(* Logix 5000 project; controller TemplateV1R0 vendor 1 type 14 code 222 rev 33.11; software revision 33.00; part 3 of 5 *)
(* tags used below, declared in another part *)
   Sts_Show_HMIControls : BOOL;   // 0 = dont show 1 = Show controls
   T_Switch_Time : TIMER[2];   // timer for valve to move from open to close or the otherway around
   ons_reset : BOOL;   // prevent continious reset
   T_Mem_Valve : TIMER[2];
(* Valve_V2, continued *)

ROUTINE Prescan   (* structured text *)
   ////////////////////////////////////////////////////////////
   //   Copyright (c)
   //------------------------------------------------------------
   //   Routine: Prescan
   //   Author: WPI\tom.reit
   //   Created: 28-11-2022
   //------------------------------------------------------------
   //   Description:
   //
   //
   //   History:
   //
   ////////////////////////////////////////////////////////////
   if T_Switch_Time[0].PRE = 0 then T_Switch_Time[0].PRE:=500; end_if;
   if T_Switch_Time[1].PRE = 0 then T_Switch_Time[1].PRE:=500; end_if;
   T_Mem_Valve[0].PRE:=50;
   T_Mem_Valve[1].PRE:=50;
   
   Sts_Show_HMIControls :=0;
   
END_ROUTINE
END_ADD_ON_INSTRUCTION

ADD_ON_INSTRUCTION WaterCircuit   (* revision 1.1, vendor WPI, ExecutePrescan *)
// Closed water circuit based on Micro820
VAR_INPUT
   Reset : BOOL; {required}   // Reset WTU C1&C2 on falling edge of reset signal
   Select_Mode : BOOL; {visible}   // 1 = Automatic 0 = Manual
   Start : BOOL; {visible}   // 0 = OFF 1 = ON
END_VAR
VAR_OUTPUT
   Temperature : REAL; {access Read Only, visible}   // Actual Temperature (c)
END_VAR
VAR_INPUT
   PID_CycleTime : DINT; {required}   // Cycle time for SSR
   PID_Kc : LREAL; {required}   // Proportional and Integral are dependent on this gain. (>= 0.0001). Increasing Kc improves response time but also increases overshoot and oscillation of the PID.
   PID_Ti : LREAL; {required}   // Time integral constant in seconds (>= 0.0001). Increasing Ti decreases the overshoot and oscillation of the PID.
   PID_Td : LREAL; {required}   // Time derivative constant in seconds (>= 0.0). When Td equals 0, there is no derivative action and PID becomes a PI controller. Increasing Td reduces the overshot and removes the oscillation of the PID controller.
   PID_FC : LREAL; {required}   // Filter constant (>= 0.0). Recommended range for FC is 0 to 20. Increasing FC smooths the response of the PID controller.
   PID_Setpoint : LREAL; {visible}   // Setpoint temperature (c)
END_VAR
VAR_OUTPUT
   PID_OUTPUT : REAL; {access Read Only, visible}   // Output PID controller (%)
END_VAR
VAR_INPUT
   PID_HandValue : LREAL; {visible}   // handvalue in % of time
   ManualStart_CP : BOOL; {visible}   // 0 = OFF 1 = ON
   ManualStart_HE : BOOL; {visible}   // 0 = OFF 1 = ON
   ManualStart_V1 : BOOL; {visible}   // 0 = OFF 1 = ON
   ManualStart_V2 : BOOL; {visible}   // 0 = OFF 1 = ON
END_VAR
VAR_OUTPUT
   ALARM_CommunicationFaulted : BOOL; {access Read Only, visible}   // Communication faulted, check IP address in MSG instruction
   ALARM_Active : BOOL; {access Read Only, visible}   // Alarm is active, outputs will NOT be activated on WTU
   ALARM_PressureFaulted : BOOL; {access Read Only, visible}   // Filling faulted
   ALARM_Overload_CirculationPump : BOOL; {access Read Only, visible}   // Overload_CirculationPump
   ALARM_Overload_Heatingelement : BOOL; {access Read Only, visible}   // Overload_Heatingelment
   ALARM_Max_TemperatureSwitch : BOOL; {access Read Only, visible}   // Max TemperatureSwitch
   ALARM_TemperatureSensorLost : BOOL; {access Read Only, visible}   // cable disconnected temperature sensor
   Sts_Communication_OK : BOOL; {access Read Only, visible}   // Communication is OK to micro820
   Sts_CirculationPump : BOOL; {access Read Only, visible}   // Status Circulationpump output
   Sts_HeatingElement : BOOL; {access Read Only, visible}   // Status Heating element output
   Sts_SolidstateRelais : BOOL; {access Read Only, visible}   // Status SSR output
   Sts_CoolingValve : BOOL; {access Read Only, visible}   // Status Cooling Valve output
   Sts_FillingValve : BOOL; {access Read Only, visible}   // Status Filling Valve output
END_VAR
VAR_IN_OUT
   Read_Element : LREAL[40]; {required}   // Dataholder
   Msg_Read : MESSAGE; {required}   // Message to read object
   Write_Element : LREAL[40]; {required}   // Dataholder
   Msg_Write : MESSAGE; {required}   // Message to read object
END_VAR
VAR_INPUT
   Enable_Communication : BOOL; {visible}   // set to true if messages can be send to micro820
   cnf_Select_Circuit : USINT;   // assign AOI to watercircuit based on: 1 = C1 2 = C2
END_VAR
VAR_OUTPUT
   HMI_Color : DINT; {access Read Only}   // 0 = off 1 = auto turned on 2 = manual control 3= no communication
END_VAR
VAR
   RefreshRate : FBD_TIMER; {access None}   // refreshrate timer
   wrk_conversion : DINT[20]; {access None}   // conversion tag to go from LREAL to DINT
   i : SINT; {access None}   // local index num
   InputStatus : DINT; {access None}   // InputStatus from Micro820
        .12   // spare
        .0   // _IO_EM_DI_00
        .1   // _IO_EM_DI_01
        .10   // _IO_EM_DI_10
        .11   // _IO_EM_DI_11
        .13   // spare
        .14   // spare
        .15   // spare
        .16   // spare
        .17   // spare
        .18   // spare
        .19   // spare
        .2   // _IO_EM_DI_02
        .20   // spare
        .21   // spare
        .22   // spare
        .23   // spare
        .24   // spare
        .25   // spare
        .26   // spare
        .27   // spare
        .28   // spare
        .29   // spare
        .3   // _IO_EM_DI_03
        .30   // spare
        .31   // spare
        .4   // _IO_EM_DI_04
        .5   // _IO_EM_DI_05
        .6   // _IO_EM_DI_06
        .7   // _IO_EM_DI_07
        .8   // _IO_EM_DI_08
        .9   // _IO_EM_DI_09
   TagName : STRING; {access Read Only}   // Contains tag name based on addon name
   HMI_Trend_MaxValue : DINT; {access Read Only}   // Trend for HMI
   HMI_Trend_MinValue : DINT; {access Read Only}   // HMI_Trend_MinValue
END_VAR

ROUTINE Logic   (* structured text *)
// Closed water circuit based on Micro820
   ////////////////////////////////////////////////////////////
   //   Copyright (c)
   //------------------------------------------------------------
   //   Routine: WaterCircuit - Logic
   //   Author: WPI\tom.reit
   //   Created: 13-3-2023
   //------------------------------------------------------------
   //   Description:
   //           Closed water circuit based on Micro820
   //
   //
   //   History:
   //
   ////////////////////////////////////////////////////////////
   RefreshRate.EN:=1;
   RefreshRate.PRE:=50;
   RefreshRate.TimerEnable:=1;
   RefreshRate.Reset:=RefreshRate.DN;
   TONR(RefreshRate);
   if RefreshRate.DN then
   	MSG(Msg_Read);																	// Message to read object. CIP datatable read.
   	MSG(Msg_Write);																	// Message to Write object. CIP datatable write.
   end_if;
   #region Message OK
   	if Msg_Read.DN AND Msg_Write.DN then
   		Sts_Communication_OK:=1;
   	end_if;
   	if NOT Enable_Communication then
   		Sts_Communication_OK:=0;
   	end_if;
   #endregion
   #region Message timeout/faulted
   	if Msg_Read.ER OR Msg_Write.ER then
   		ALARM_CommunicationFaulted:=1;
   		Sts_Communication_OK:=0;
   	else
   		ALARM_CommunicationFaulted:=0;
   	end_if;
   	if Reset AND (Msg_Read.ER OR Msg_Write.ER)  then
   		Msg_Read.Flags			:=0;	// reset Message instruction
   		Msg_Write.Flags			:=0;	// reset Message instruction
   	end_if;
   #endregion
   for i := 0 to 19 do
   	wrk_conversion[i]:=0;// clear old data
   end_for;
   wrk_conversion[0].0			:=		Reset;						// Micro820 tag: HMI_I_Reset
   
   /* Prevent wrong user input */
   if cnf_Select_Circuit > 2 then cnf_Select_Circuit:=2; end_if;
   if cnf_Select_Circuit < 1 then cnf_Select_Circuit:=1; end_if;
   
   #region Convert IO from Micro820 to local
   	wrk_conversion[18]				:=		Read_Element[18];	// InputStatus
   	InputStatus						:= 		wrk_conversion[18];
   	wrk_conversion[19]				:=		Read_Element[19];	// OutputStatus
   #endregion
   if Enable_Communication then
   	#region data
   		#region Convert InputData to LREAL
   			wrk_conversion[1].0			:=		Select_Mode;				// Micro820 tag: HMI_I_C1_Select_Mode
   			wrk_conversion[2].0			:=		Start;					// Micro820 tag: HMI_I_StartC1
   			wrk_conversion[3].0			:=		ManualStart_CP;			// Micro820 tag: HMI_I_C1_ManualStart_CP
   			wrk_conversion[4].0			:=		ManualStart_HE;			// Micro820 tag: HMI_I_C1_ManualStart_HE
   			wrk_conversion[5].0			:=		ManualStart_V1;			// Micro820 tag: HMI_I_C1_ManualStart_V1
   			wrk_conversion[6].0			:=		ManualStart_V2;			// Micro820 tag: HMI_I_C1_ManualStart_V2
   			// IS ALLREADY A REAL, DOESNT NEED CONVERSION! 					// Micro820 tag: HMI_I_C1_Kc
   			// IS ALLREADY A REAL, DOESNT NEED CONVERSION! 					// Micro820 tag: HMI_I_C1_Ti
   			// IS ALLREADY A REAL, DOESNT NEED CONVERSION! 					// Micro820 tag: HMI_I_C1_Td
   			// IS ALLREADY A REAL, DOESNT NEED CONVERSION! 					// Micro820 tag: HMI_I_C1_FC
   			// IS ALLREADY A REAL, DOESNT NEED CONVERSION! 					// Micro820 tag: HMI_I_C1_PID_Setpoint
   			// IS ALLREADY A REAL, DOESNT NEED CONVERSION!					// Micro820 tag: HMI_I_C1_PID_HandValue
   			wrk_conversion[13]			:=		PID_CycleTime;			// Micro820 tag: HMI_I_C1_PID_CycleTime
   		/* set data for micro820 tag */
   		Write_Element[00]:=wrk_conversion[00];
   		Write_Element[01]:=wrk_conversion[01];
   		Write_Element[02]:=wrk_conversion[02];
   		Write_Element[03]:=wrk_conversion[03];
   		Write_Element[04]:=wrk_conversion[04];
   		Write_Element[05]:=wrk_conversion[05];
   		Write_Element[06]:=wrk_conversion[06];
   		Write_Element[07]:=PID_Kc;
   		Write_Element[08]:=PID_Ti;
   		Write_Element[09]:=PID_Td;
   		Write_Element[10]:=PID_FC;
   		Write_Element[11]:=PID_Setpoint;
   		Write_Element[12]:=PID_HandValue;
   		Write_Element[13]:=wrk_conversion[13];
   		#endregion
   		#region OutputData
   			Temperature						:=		Read_Element[0];
   			PID_OUTPUT						:=		Read_Element[1];
   
   			wrk_conversion[2]				:=		Read_Element[2];
   			ALARM_PressureFaulted			:=		wrk_conversion[2].0;
   
   			wrk_conversion[3]				:=		Read_Element[3];
   			ALARM_Overload_CirculationPump	:=		wrk_conversion[3].0;
   
   			wrk_conversion[4]				:=		Read_Element[4];
   			ALARM_Overload_Heatingelement	:=		wrk_conversion[4].0;
   
   			wrk_conversion[5]				:=		Read_Element[5];
   			ALARM_Max_TemperatureSwitch		:=		wrk_conversion[5].0;
   
   			wrk_conversion[6]				:=		Read_Element[6];
   			ALARM_TemperatureSensorLost		:=		wrk_conversion[6].0;
   
   			wrk_conversion[7]				:=		Read_Element[7];
   			ALARM_Active					:=		wrk_conversion[7].0;
   
   			if cnf_Select_Circuit = 1 then
   				Sts_CirculationPump				:=		wrk_conversion[19].0;
   				Sts_HeatingElement				:=		wrk_conversion[19].1;
   				Sts_SolidstateRelais			:=		wrk_conversion[19].2;
   				Sts_CoolingValve				:=		wrk_conversion[19].3;
   				Sts_FillingValve				:=		wrk_conversion[19].4;
   			elsif cnf_Select_Circuit = 2 then
   				Sts_CirculationPump				:=		wrk_conversion[19].5;
   				Sts_HeatingElement				:=		wrk_conversion[19].6;
   				Sts_SolidstateRelais			:=		wrk_conversion[19].7;
   				Sts_CoolingValve				:=		wrk_conversion[19].8;
   				Sts_FillingValve				:=		wrk_conversion[19].9;
   			end_if;
   		#endregion
   	#endregion
   end_if;
   #region HMI data visuals
   	if 	(Enable_Communication AND Sts_Communication_OK )  AND Select_Mode AND NOT Start then			// Auto - Turned off
   		HMI_Color:=0;
   	elsif (Enable_Communication AND Sts_Communication_OK )  AND Select_Mode AND Start then				// Auto - Turned on
   		HMI_Color:=1;
   	elsif (Enable_Communication AND Sts_Communication_OK )  AND NOT Select_Mode  then					// Manual - controlled manually
   		HMI_Color:=2;
   	elsif (Enable_Communication AND NOT Sts_Communication_OK ) then										// No connection
   		HMI_Color:=0;
   	elsif NOT Enable_Communication then																	// No connection
   		HMI_Color:=3;
   	end_if;
   	gsv(AddOnInstructionDefinition,THIS,Name,TagName);
   	if HMI_Trend_MaxValue=0 AND HMI_Trend_MinValue=0 then HMI_Trend_MaxValue:=100;HMI_Trend_MinValue:=0; end_if;
   #endregion
END_ROUTINE

ROUTINE Prescan   (* structured text *)
   ////////////////////////////////////////////////////////////
   //   Copyright (c)
   //------------------------------------------------------------
   //   Routine: Prescan
   //   Author: WPI\tom.reit
   //   Created: 15-3-2023
   //------------------------------------------------------------
   //   Description:
   //
   //
   //   History:
   //
   ////////////////////////////////////////////////////////////
   Enable_Communication:=1;
END_ROUTINE
END_ADD_ON_INSTRUCTION

VAR_GLOBAL   (* controller tags *)
   SafetyZone1_Unit1_Reset : BOOL;
END_VAR

PROGRAM MainProgram   (* main routine MainRoutine *)

ROUTINE MainRoutine   (* ladder *)
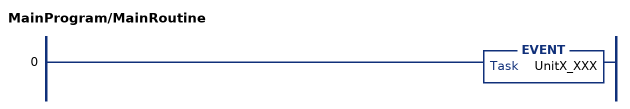
   0: EVENT(UnitX_XXX);
END_ROUTINE
END_PROGRAM

PROGRAM SafetyProgram   (* main routine MainRoutine, safety *)

ROUTINE MainRoutine   (* ladder *)
END_ROUTINE
END_PROGRAM

PROGRAM UnitX_EMXXX   (* main routine Main *)
VAR
   Alarm : AlarmGenerator[10] := ([1].Alarm_ID := 1, [2].Alarm_ID := 2, [3].Alarm_ID := 3, [4].Alarm_ID := 4, [5].Alarm_ID := 5, [6].Alarm_ID := 6, [7].Alarm_ID := 7, [8].Alarm_ID := 8, [9].Alarm_ID := 9);
   AlarmText : STRING[10] := ([1] := '| Unit4_Batter_EM01_Depositor | X-axis faulted | ', [2] := '| Unit4_Batter_EM01_Depositor | Y-axis faulted |', [3] := '| Unit4_Batter_EM01_Depositor | Z-axis faulted |', [4] := '| Unit4_Batter_EM01_Depositor | Manifold ColorInjected-axis faulted |', [5] := '| Unit4_Batter_EM01_Depositor | No Color Manifold-axis faulted |', [6] := '| Unit4_Batter_EM01_Depositor | Overload servo drives |', [7] := '| Unit4_Batter_EM01_Depositor | X,Y,Z Motion faulted |', [8] := '| Unit4_Batter_EM01_Depositor | Manifold Motion faulted |', [9] := '| Unit1_Sander_EM01_Elende |');
   wrk_mode_Select : DINT := 1;   // mode select for case
   wrk_StartNum : DINT := 100;   // StartStateModelNum
   wrk_state_Select : DINT := 9;   // select correct prog
END_VAR

ROUTINE _EP_00_Selector   (* structured text *)
   ////////////////////////////////////////////////////////////
   //   Copyright (c)
   //------------------------------------------------------------
   //   Routine: _EP_00_Selector
   //   Author: WPI\tom.reit
   //   Created: 11-11-2022
   //------------------------------------------------------------
   //   Description:
   //
   //
   //   History:
   //
   ////////////////////////////////////////////////////////////
   if 		Unit.Sts_Production 	then	wrk_mode_Select:=1;
   elsif 	Unit.Sts_Maintenance 	then	wrk_mode_Select:=2;
   elsif 	Unit.Sts_Manual 		then	wrk_mode_Select:=3;
   elsif 	Unit.Sts_Cleaning 		then	wrk_mode_Select:=4;
   elsif 	Unit.Sts_MES 			then	wrk_mode_Select:=5;
   elsif 	Unit.Sts_SemiAutomatic 	then	wrk_mode_Select:=6;
   end_if;
   #region Set case state non active states
   	if 		Unit.Sts_Aborted 		then	wrk_state_Select:=9;
   	elsif 	Unit.Sts_Stopped		then	wrk_state_Select:=2;
   	elsif   Unit.Sts_Idle			then	wrk_state_Select:=4;
   	elsif 	Unit.Sts_Execute		then	wrk_state_Select:=6;
   	elsif 	Unit.Sts_Held			then	wrk_state_Select:=11;
   	elsif 	Unit.Sts_Suspended		then	wrk_state_Select:=5;
   	elsif   Unit.Sts_Complete		then	wrk_state_Select:=17;
   	end_if;
   #endregion
   #region Set case state
   	if 		Unit.Sts_Production AND Unit.Sts_Aborting 		then	wrk_state_Select:=8;
   	elsif 	Unit.Sts_Production AND Unit.Sts_Clearing		then	wrk_state_Select:=1;
   	elsif 	Unit.Sts_Production AND Unit.Sts_Stopping		then	wrk_state_Select:=7;
   	elsif 	Unit.Sts_Production	AND Unit.Sts_Resetting		then	wrk_state_Select:=15;
   	elsif 	Unit.Sts_Production AND Unit.Sts_Starting		then	wrk_state_Select:=3;
   	elsif 	Unit.Sts_Production AND Unit.Sts_Holding		then	wrk_state_Select:=10;
   	elsif 	Unit.Sts_Production AND Unit.Sts_Unholding		then	wrk_state_Select:=12;
   	elsif 	Unit.Sts_Production AND Unit.Sts_Suspending		then	wrk_state_Select:=13;
   	elsif 	Unit.Sts_Production AND Unit.Sts_Unsuspending	then	wrk_state_Select:=14;
   	elsif 	Unit.Sts_Production AND Unit.Sts_Completing		then	wrk_state_Select:=16;
   	end_if;
   #endregion
   #region Set case state
   	if 		Unit.Sts_Maintenance AND Unit.Sts_Aborting 		then	wrk_state_Select:=8;
   	elsif 	Unit.Sts_Maintenance AND Unit.Sts_Clearing		then	wrk_state_Select:=1;
   	elsif 	Unit.Sts_Maintenance AND Unit.Sts_Stopping		then	wrk_state_Select:=7;
   	elsif 	Unit.Sts_Maintenance AND Unit.Sts_Resetting		then	wrk_state_Select:=15;
   	elsif 	Unit.Sts_Maintenance AND Unit.Sts_Starting		then	wrk_state_Select:=3;
   	elsif 	Unit.Sts_Maintenance AND Unit.Sts_Holding		then	wrk_state_Select:=10;
   	elsif 	Unit.Sts_Maintenance AND Unit.Sts_Unholding		then	wrk_state_Select:=12;
   	elsif 	Unit.Sts_Maintenance AND Unit.Sts_Suspending	then	wrk_state_Select:=13;
   	elsif 	Unit.Sts_Maintenance AND Unit.Sts_Unsuspending	then	wrk_state_Select:=14;
   	elsif 	Unit.Sts_Maintenance AND Unit.Sts_Completing	then	wrk_state_Select:=16;
   	end_if;
   #endregion
   #region Set case state
   	if 		Unit.Sts_Manual AND Unit.Sts_Aborting 		then	wrk_state_Select:=8;
   	elsif 	Unit.Sts_Manual AND Unit.Sts_Clearing		then	wrk_state_Select:=1;
   	elsif 	Unit.Sts_Manual AND Unit.Sts_Stopping		then	wrk_state_Select:=7;
   	elsif 	Unit.Sts_Manual	AND Unit.Sts_Resetting		then	wrk_state_Select:=15;
   	elsif 	Unit.Sts_Manual AND Unit.Sts_Starting		then	wrk_state_Select:=3;
   	elsif 	Unit.Sts_Manual AND Unit.Sts_Holding		then	wrk_state_Select:=10;
   	elsif 	Unit.Sts_Manual AND Unit.Sts_Unholding		then	wrk_state_Select:=12;
   	elsif 	Unit.Sts_Manual AND Unit.Sts_Suspending		then	wrk_state_Select:=13;
   	elsif 	Unit.Sts_Manual AND Unit.Sts_Unsuspending	then	wrk_state_Select:=14;
   	elsif 	Unit.Sts_Manual AND Unit.Sts_Completing		then	wrk_state_Select:=16;
   	end_if;
   #endregion
   #region Set case state
   	if 		Unit.Sts_Cleaning AND Unit.Sts_Aborting 	then	wrk_state_Select:=8;
   	elsif 	Unit.Sts_Cleaning AND Unit.Sts_Clearing		then	wrk_state_Select:=1;
   	elsif 	Unit.Sts_Cleaning AND Unit.Sts_Stopping		then	wrk_state_Select:=7;
   	elsif 	Unit.Sts_Cleaning AND Unit.Sts_Resetting	then	wrk_state_Select:=15;
   	elsif 	Unit.Sts_Cleaning AND Unit.Sts_Starting		then	wrk_state_Select:=3;
   	elsif 	Unit.Sts_Cleaning AND Unit.Sts_Holding		then	wrk_state_Select:=10;
   	elsif 	Unit.Sts_Cleaning AND Unit.Sts_Unholding	then	wrk_state_Select:=12;
   	elsif 	Unit.Sts_Cleaning AND Unit.Sts_Suspending	then	wrk_state_Select:=13;
   	elsif 	Unit.Sts_Cleaning AND Unit.Sts_Unsuspending	then	wrk_state_Select:=14;
   	elsif 	Unit.Sts_Cleaning AND Unit.Sts_Completing	then	wrk_state_Select:=16;
   	end_if;
   #endregion
   #region Set case state
   	if 		Unit.Sts_MES AND Unit.Sts_Aborting 		then	wrk_state_Select:=8;
   	elsif 	Unit.Sts_MES AND Unit.Sts_Clearing		then	wrk_state_Select:=1;
   	elsif 	Unit.Sts_MES AND Unit.Sts_Stopping		then	wrk_state_Select:=7;
   	elsif 	Unit.Sts_MES AND Unit.Sts_Resetting		then	wrk_state_Select:=15;
   	elsif 	Unit.Sts_MES AND Unit.Sts_Starting		then	wrk_state_Select:=3;
   	elsif 	Unit.Sts_MES AND Unit.Sts_Holding		then	wrk_state_Select:=10;
   	elsif 	Unit.Sts_MES AND Unit.Sts_Unholding		then	wrk_state_Select:=12;
   	elsif 	Unit.Sts_MES AND Unit.Sts_Suspending	then	wrk_state_Select:=13;
   	elsif 	Unit.Sts_MES AND Unit.Sts_Unsuspending	then	wrk_state_Select:=14;
   	elsif 	Unit.Sts_MES AND Unit.Sts_Completing	then	wrk_state_Select:=16;
   	end_if;
   #endregion
   #region Set case state
   	if 		Unit.Sts_SemiAutomatic AND Unit.Sts_Aborting 		then	wrk_state_Select:=8;
   	elsif 	Unit.Sts_SemiAutomatic AND Unit.Sts_Clearing		then	wrk_state_Select:=1;
   	elsif 	Unit.Sts_SemiAutomatic AND Unit.Sts_Stopping		then	wrk_state_Select:=7;
   	elsif 	Unit.Sts_SemiAutomatic	AND Unit.Sts_Resetting		then	wrk_state_Select:=15;
   	elsif 	Unit.Sts_SemiAutomatic AND Unit.Sts_Starting		then	wrk_state_Select:=3;
   	elsif 	Unit.Sts_SemiAutomatic AND Unit.Sts_Holding			then	wrk_state_Select:=10;
   	elsif 	Unit.Sts_SemiAutomatic AND Unit.Sts_Unholding		then	wrk_state_Select:=12;
   	elsif 	Unit.Sts_SemiAutomatic AND Unit.Sts_Suspending		then	wrk_state_Select:=13;
   	elsif 	Unit.Sts_SemiAutomatic AND Unit.Sts_Unsuspending	then	wrk_state_Select:=14;
   	elsif 	Unit.Sts_SemiAutomatic AND Unit.Sts_Completing		then	wrk_state_Select:=16;
   	end_if;
   #endregion
   
   
   EquipmentModule.Request_SC.ons_Reset.InputBit:=Unit.Sts_MachineFaulted OR EquipmentModule.Reset_Signal;
   OSRI(EquipmentModule.Request_SC.ons_Reset);
   if EquipmentModule.Request_SC.ons_Reset.OutputBit then
   	EquipmentModule.EP_SEQ.Holding		:=0;
   	EquipmentModule.EP_SEQ.Starting		:=0;
   	EquipmentModule.EP_SEQ.Suspending	:=0;
   	EquipmentModule.EP_SEQ.Unholding	:=0;
   	EquipmentModule.EP_SEQ.Unsuspending	:=0;
   end_if;
   
   if EquipmentModule.Force_Stop OR EquipmentModule.Force_Abort then EquipmentModule.Faulted:=1; else EquipmentModule.Faulted:=0; end_if;
   case wrk_mode_Select of
   	1:																	/* Production(automatic) */
   		wrk_StartNum:=100;
   		case wrk_state_Select of
   			1: 	JSR(_EP_01_Clearing); 		if EquipmentModule.EP_SEQ.Clearing		=0 then EquipmentModule.EP_SEQ.Clearing		:=wrk_StartNum; 	end_if;
   			3: 	JSR(_EP_03_Starting);		if EquipmentModule.EP_SEQ.Starting		=0 then EquipmentModule.EP_SEQ.Starting		:=wrk_StartNum; 	end_if;
   			6: 	JSR(_EP_06_Execute);
   			7: 	JSR(_EP_07_Stopping);		if EquipmentModule.EP_SEQ.Stopping		=0 then EquipmentModule.EP_SEQ.Stopping		:=wrk_StartNum; 	end_if;
   			8: 	JSR(_EP_08_Aborting); 		if EquipmentModule.EP_SEQ.Aborting		=0 then EquipmentModule.EP_SEQ.Aborting		:=wrk_StartNum; 	end_if;
   			10: JSR(_EP_10_Holding);		if EquipmentModule.EP_SEQ.Holding		=0 then EquipmentModule.EP_SEQ.Holding		:=wrk_StartNum; 	end_if;
   			12:	JSR(_EP_12_Unholding);		if EquipmentModule.EP_SEQ.Unholding		=0 then EquipmentModule.EP_SEQ.Unholding	:=wrk_StartNum; 	end_if;
   			13:	JSR(_EP_13_Suspending);		if EquipmentModule.EP_SEQ.Suspending	=0 then EquipmentModule.EP_SEQ.Suspending	:=wrk_StartNum; 	end_if;
   			14:	JSR(_EP_14_Unsuspending);	if EquipmentModule.EP_SEQ.Unsuspending	=0 then EquipmentModule.EP_SEQ.Unsuspending	:=wrk_StartNum; 	end_if;
   			15:	JSR(_EP_15_Resetting);		if EquipmentModule.EP_SEQ.Resetting		=0 then EquipmentModule.EP_SEQ.Resetting	:=wrk_StartNum; 	end_if;
   			16:	JSR(_EP_16_Completing);		if EquipmentModule.EP_SEQ.Completing	=0 then EquipmentModule.EP_SEQ.Completing	:=wrk_StartNum; 	end_if;
   			else
   		end_case;
   	2:																	/* Maintenance */
   		wrk_StartNum:=200;
   		case wrk_state_Select of
   			1: 	JSR(_EP_01_Clearing); 		if EquipmentModule.EP_SEQ.Clearing		=0 then EquipmentModule.EP_SEQ.Clearing		:=wrk_StartNum; 	end_if;
   			3: 	JSR(_EP_03_Starting);		if EquipmentModule.EP_SEQ.Starting		=0 then EquipmentModule.EP_SEQ.Starting		:=wrk_StartNum; 	end_if;
   			6: 	JSR(_EP_06_Execute);
   			7: 	JSR(_EP_07_Stopping);		if EquipmentModule.EP_SEQ.Stopping		=0 then EquipmentModule.EP_SEQ.Stopping		:=wrk_StartNum; 	end_if;
   			8: 	JSR(_EP_08_Aborting); 		if EquipmentModule.EP_SEQ.Aborting		=0 then EquipmentModule.EP_SEQ.Aborting		:=wrk_StartNum; 	end_if;
   			10: JSR(_EP_10_Holding);		if EquipmentModule.EP_SEQ.Holding		=0 then EquipmentModule.EP_SEQ.Holding		:=wrk_StartNum; 	end_if;
   			12:	JSR(_EP_12_Unholding);		if EquipmentModule.EP_SEQ.Unholding		=0 then EquipmentModule.EP_SEQ.Unholding	:=wrk_StartNum; 	end_if;
   			13:	JSR(_EP_13_Suspending);		if EquipmentModule.EP_SEQ.Suspending	=0 then EquipmentModule.EP_SEQ.Suspending	:=wrk_StartNum; 	end_if;
   			14:	JSR(_EP_14_Unsuspending);	if EquipmentModule.EP_SEQ.Unsuspending	=0 then EquipmentModule.EP_SEQ.Unsuspending	:=wrk_StartNum; 	end_if;
   			15:	JSR(_EP_15_Resetting);		if EquipmentModule.EP_SEQ.Resetting		=0 then EquipmentModule.EP_SEQ.Resetting	:=wrk_StartNum; 	end_if;
   			16:	JSR(_EP_16_Completing);		if EquipmentModule.EP_SEQ.Completing	=0 then EquipmentModule.EP_SEQ.Completing	:=wrk_StartNum; 	end_if;
   			else
   		end_case;
   	3:																	/* Manual */
   		wrk_StartNum:=300;
   		case wrk_state_Select of
   			1: 	JSR(_EP_01_Clearing); 		if EquipmentModule.EP_SEQ.Clearing		=0 then EquipmentModule.EP_SEQ.Clearing		:=wrk_StartNum; 	end_if;
   			3: 	JSR(_EP_03_Starting);		if EquipmentModule.EP_SEQ.Starting		=0 then EquipmentModule.EP_SEQ.Starting		:=wrk_StartNum; 	end_if;
   			6: 	JSR(_EP_06_Execute);
   			7: 	JSR(_EP_07_Stopping);		if EquipmentModule.EP_SEQ.Stopping		=0 then EquipmentModule.EP_SEQ.Stopping		:=wrk_StartNum; 	end_if;
   			8: 	JSR(_EP_08_Aborting); 		if EquipmentModule.EP_SEQ.Aborting		=0 then EquipmentModule.EP_SEQ.Aborting		:=wrk_StartNum; 	end_if;
   			10: JSR(_EP_10_Holding);		if EquipmentModule.EP_SEQ.Holding		=0 then EquipmentModule.EP_SEQ.Holding		:=wrk_StartNum; 	end_if;
   			12:	JSR(_EP_12_Unholding);		if EquipmentModule.EP_SEQ.Unholding		=0 then EquipmentModule.EP_SEQ.Unholding	:=wrk_StartNum; 	end_if;
   			13:	JSR(_EP_13_Suspending);		if EquipmentModule.EP_SEQ.Suspending	=0 then EquipmentModule.EP_SEQ.Suspending	:=wrk_StartNum; 	end_if;
   			14:	JSR(_EP_14_Unsuspending);	if EquipmentModule.EP_SEQ.Unsuspending	=0 then EquipmentModule.EP_SEQ.Unsuspending	:=wrk_StartNum; 	end_if;
   			15:	JSR(_EP_15_Resetting);		if EquipmentModule.EP_SEQ.Resetting		=0 then EquipmentModule.EP_SEQ.Resetting	:=wrk_StartNum; 	end_if;
   			16:	JSR(_EP_16_Completing);		if EquipmentModule.EP_SEQ.Completing	=0 then EquipmentModule.EP_SEQ.Completing	:=wrk_StartNum; 	end_if;
   			else
   		end_case;
   	4:																	/* Cleaning */
   		wrk_StartNum:=400;
   		case wrk_state_Select of
   			1: 	JSR(_EP_01_Clearing); 		if EquipmentModule.EP_SEQ.Clearing		=0 then EquipmentModule.EP_SEQ.Clearing		:=wrk_StartNum; 	end_if;
   			3: 	JSR(_EP_03_Starting);		if EquipmentModule.EP_SEQ.Starting		=0 then EquipmentModule.EP_SEQ.Starting		:=wrk_StartNum; 	end_if;
   			6: 	JSR(_EP_06_Execute);
   			7: 	JSR(_EP_07_Stopping);		if EquipmentModule.EP_SEQ.Stopping		=0 then EquipmentModule.EP_SEQ.Stopping		:=wrk_StartNum; 	end_if;
   			8: 	JSR(_EP_08_Aborting); 		if EquipmentModule.EP_SEQ.Aborting		=0 then EquipmentModule.EP_SEQ.Aborting		:=wrk_StartNum; 	end_if;
   			10: JSR(_EP_10_Holding);		if EquipmentModule.EP_SEQ.Holding		=0 then EquipmentModule.EP_SEQ.Holding		:=wrk_StartNum; 	end_if;
   			12:	JSR(_EP_12_Unholding);		if EquipmentModule.EP_SEQ.Unholding		=0 then EquipmentModule.EP_SEQ.Unholding	:=wrk_StartNum; 	end_if;
   			13:	JSR(_EP_13_Suspending);		if EquipmentModule.EP_SEQ.Suspending	=0 then EquipmentModule.EP_SEQ.Suspending	:=wrk_StartNum; 	end_if;
   			14:	JSR(_EP_14_Unsuspending);	if EquipmentModule.EP_SEQ.Unsuspending	=0 then EquipmentModule.EP_SEQ.Unsuspending	:=wrk_StartNum; 	end_if;
   			15:	JSR(_EP_15_Resetting);		if EquipmentModule.EP_SEQ.Resetting		=0 then EquipmentModule.EP_SEQ.Resetting	:=wrk_StartNum; 	end_if;
   			16:	JSR(_EP_16_Completing);		if EquipmentModule.EP_SEQ.Completing	=0 then EquipmentModule.EP_SEQ.Completing	:=wrk_StartNum; 	end_if;
   			else
   		end_case;
   	5:																	/* MES */
   		wrk_StartNum:=500;
   		case wrk_state_Select of
   			1: 	JSR(_EP_01_Clearing); 		if EquipmentModule.EP_SEQ.Clearing		=0 then EquipmentModule.EP_SEQ.Clearing		:=wrk_StartNum; 	end_if;
   			3: 	JSR(_EP_03_Starting);		if EquipmentModule.EP_SEQ.Starting		=0 then EquipmentModule.EP_SEQ.Starting		:=wrk_StartNum; 	end_if;
   			6: 	JSR(_EP_06_Execute);
   			7: 	JSR(_EP_07_Stopping);		if EquipmentModule.EP_SEQ.Stopping		=0 then EquipmentModule.EP_SEQ.Stopping		:=wrk_StartNum; 	end_if;
   			8: 	JSR(_EP_08_Aborting); 		if EquipmentModule.EP_SEQ.Aborting		=0 then EquipmentModule.EP_SEQ.Aborting		:=wrk_StartNum; 	end_if;
   			10: JSR(_EP_10_Holding);		if EquipmentModule.EP_SEQ.Holding		=0 then EquipmentModule.EP_SEQ.Holding		:=wrk_StartNum; 	end_if;
   			12:	JSR(_EP_12_Unholding);		if EquipmentModule.EP_SEQ.Unholding		=0 then EquipmentModule.EP_SEQ.Unholding	:=wrk_StartNum; 	end_if;
   			13:	JSR(_EP_13_Suspending);		if EquipmentModule.EP_SEQ.Suspending	=0 then EquipmentModule.EP_SEQ.Suspending	:=wrk_StartNum; 	end_if;
   			14:	JSR(_EP_14_Unsuspending);	if EquipmentModule.EP_SEQ.Unsuspending	=0 then EquipmentModule.EP_SEQ.Unsuspending	:=wrk_StartNum; 	end_if;
   			15:	JSR(_EP_15_Resetting);		if EquipmentModule.EP_SEQ.Resetting		=0 then EquipmentModule.EP_SEQ.Resetting	:=wrk_StartNum; 	end_if;
   			16:	JSR(_EP_16_Completing);		if EquipmentModule.EP_SEQ.Completing	=0 then EquipmentModule.EP_SEQ.Completing	:=wrk_StartNum; 	end_if;
   			else
   		end_case;
   	6:																	/* semiautomatic */
   		wrk_StartNum:=600;
   		case wrk_state_Select of
   			1: 	JSR(_EP_01_Clearing); 		if EquipmentModule.EP_SEQ.Clearing		=0 then EquipmentModule.EP_SEQ.Clearing		:=wrk_StartNum; 	end_if;
   			3: 	JSR(_EP_03_Starting);		if EquipmentModule.EP_SEQ.Starting		=0 then EquipmentModule.EP_SEQ.Starting		:=wrk_StartNum; 	end_if;
   			6: 	JSR(_EP_06_Execute);
   			7: 	JSR(_EP_07_Stopping);		if EquipmentModule.EP_SEQ.Stopping		=0 then EquipmentModule.EP_SEQ.Stopping		:=wrk_StartNum; 	end_if;
   			8: 	JSR(_EP_08_Aborting); 		if EquipmentModule.EP_SEQ.Aborting		=0 then EquipmentModule.EP_SEQ.Aborting		:=wrk_StartNum; 	end_if;
   			10: JSR(_EP_10_Holding);		if EquipmentModule.EP_SEQ.Holding		=0 then EquipmentModule.EP_SEQ.Holding		:=wrk_StartNum; 	end_if;
   			12:	JSR(_EP_12_Unholding);		if EquipmentModule.EP_SEQ.Unholding		=0 then EquipmentModule.EP_SEQ.Unholding	:=wrk_StartNum; 	end_if;
   			13:	JSR(_EP_13_Suspending);		if EquipmentModule.EP_SEQ.Suspending	=0 then EquipmentModule.EP_SEQ.Suspending	:=wrk_StartNum; 	end_if;
   			14:	JSR(_EP_14_Unsuspending);	if EquipmentModule.EP_SEQ.Unsuspending	=0 then EquipmentModule.EP_SEQ.Unsuspending	:=wrk_StartNum; 	end_if;
   			15:	JSR(_EP_15_Resetting);		if EquipmentModule.EP_SEQ.Resetting		=0 then EquipmentModule.EP_SEQ.Resetting	:=wrk_StartNum; 	end_if;
   			16:	JSR(_EP_16_Completing);		if EquipmentModule.EP_SEQ.Completing	=0 then EquipmentModule.EP_SEQ.Completing	:=wrk_StartNum; 	end_if;
   			else
   		end_case;
   	else
   		wrk_mode_Select:=1;
   end_case;
   
   													/* Reset SC signals once machine is next state */
   if Unit.Sts_Aborted 	AND EquipmentModule.Request_SC.Aborting_to_Aborted 		then EquipmentModule.Request_SC.Aborting_to_Aborted			:=0; 	end_if;
   if Unit.Sts_Complete 	AND EquipmentModule.Request_SC.Completing_to_Completed 	then EquipmentModule.Request_SC.Completing_to_Completed		:=0; 	end_if;
   if Unit.Sts_Execute 	AND EquipmentModule.Request_SC.Starting_to_Execute 		then EquipmentModule.Request_SC.Starting_to_Execute			:=0; 	end_if;
   if Unit.Sts_Complete 	AND EquipmentModule.Request_SC.Execute_to_Completing 	then EquipmentModule.Request_SC.Execute_to_Completing		:=0; 	end_if;
   if Unit.Sts_Execute 	AND EquipmentModule.Request_SC.Unholding_to_Execute 	then EquipmentModule.Request_SC.Unholding_to_Execute		:=0; 	end_if;
   if Unit.Sts_Execute 	AND EquipmentModule.Request_SC.Unsuspending_to_Execute 	then EquipmentModule.Request_SC.Unsuspending_to_Execute		:=0; 	end_if;
   if Unit.Sts_Held 		AND EquipmentModule.Request_SC.Holding_to_Held 			then EquipmentModule.Request_SC.Holding_to_Held				:=0; 	end_if;
   if Unit.Sts_Idle 		AND EquipmentModule.Request_SC.Resetting_to_Idle 		then EquipmentModule.Request_SC.Resetting_to_Idle			:=0; 	end_if;
   if Unit.Sts_Stopped 	AND EquipmentModule.Request_SC.Clearing_to_Stopped 		then EquipmentModule.Request_SC.Clearing_to_Stopped 		:=0; 	end_if;
   if Unit.Sts_Stopped 	AND EquipmentModule.Request_SC.Stopping_to_Stopped 		then EquipmentModule.Request_SC.Stopping_to_Stopped			:=0; 	end_if;
   if Unit.Sts_Suspended 	AND EquipmentModule.Request_SC.Suspending_to_Suspended 	then EquipmentModule.Request_SC.Suspending_to_Suspended		:=0; 	end_if;
   
   													/* Reset SEQ once machine is next state */
   if Unit.Sts_Aborted 	AND		EquipmentModule.EP_SEQ.Aborting<>0		then EquipmentModule.EP_SEQ.Aborting	:=0; end_if;
   if Unit.Sts_Stopped 	AND		EquipmentModule.EP_SEQ.Clearing<>0		then EquipmentModule.EP_SEQ.Clearing	:=0; end_if;
   if Unit.Sts_Stopped 	AND		EquipmentModule.EP_SEQ.Stopping<>0		then EquipmentModule.EP_SEQ.Stopping	:=0; end_if;
   if Unit.Sts_Idle 		AND		EquipmentModule.EP_SEQ.Resetting<>0		then EquipmentModule.EP_SEQ.Resetting	:=0; end_if;
   if Unit.Sts_Execute 	AND		EquipmentModule.EP_SEQ.Starting<>0		then EquipmentModule.EP_SEQ.Starting	:=0; end_if;
   if Unit.Sts_Execute 	AND		EquipmentModule.EP_SEQ.Unholding<>0		then EquipmentModule.EP_SEQ.Unholding	:=0; end_if;
   if Unit.Sts_Execute 	AND		EquipmentModule.EP_SEQ.Unsuspending<>0	then EquipmentModule.EP_SEQ.Unsuspending:=0; end_if;
   if Unit.Sts_Complete 	AND		EquipmentModule.EP_SEQ.Completing<>0	then EquipmentModule.EP_SEQ.Completing	:=0; end_if;
   if Unit.Sts_Held 		AND		EquipmentModule.EP_SEQ.Holding<>0		then EquipmentModule.EP_SEQ.Holding		:=0; end_if;
   if Unit.Sts_Suspended	AND		EquipmentModule.EP_SEQ.Suspending<>0	then EquipmentModule.EP_SEQ.Suspending	:=0; end_if;
   
   
   
   
   
   #region AlarmFeedback to Unit
   	Alarm[1].Alarm_ID:=1;
   	Alarm[2].Alarm_ID:=2;
   	Alarm[3].Alarm_ID:=3;
   	Alarm[4].Alarm_ID:=4;
   	Alarm[5].Alarm_ID:=5;
   	Alarm[6].Alarm_ID:=6;
   	Alarm[7].Alarm_ID:=7;
   	Alarm[8].Alarm_ID:=8;
   	Alarm[9].Alarm_ID:=9;
   	AlarmGenerator(Alarm[1],EquipmentModule,AlarmText[1]);
   	AlarmGenerator(Alarm[2],EquipmentModule,AlarmText[2]);
   	AlarmGenerator(Alarm[3],EquipmentModule,AlarmText[3]);
   	AlarmGenerator(Alarm[4],EquipmentModule,AlarmText[4]);
   	AlarmGenerator(Alarm[5],EquipmentModule,AlarmText[5]);
   	AlarmGenerator(Alarm[6],EquipmentModule,AlarmText[6]);
   	AlarmGenerator(Alarm[7],EquipmentModule,AlarmText[7]);
   	AlarmGenerator(Alarm[8],EquipmentModule,AlarmText[8]);
   	AlarmGenerator(Alarm[9],EquipmentModule,AlarmText[9]);
   #endregion
END_ROUTINE

ROUTINE _EP_01_Clearing   (* ladder *)
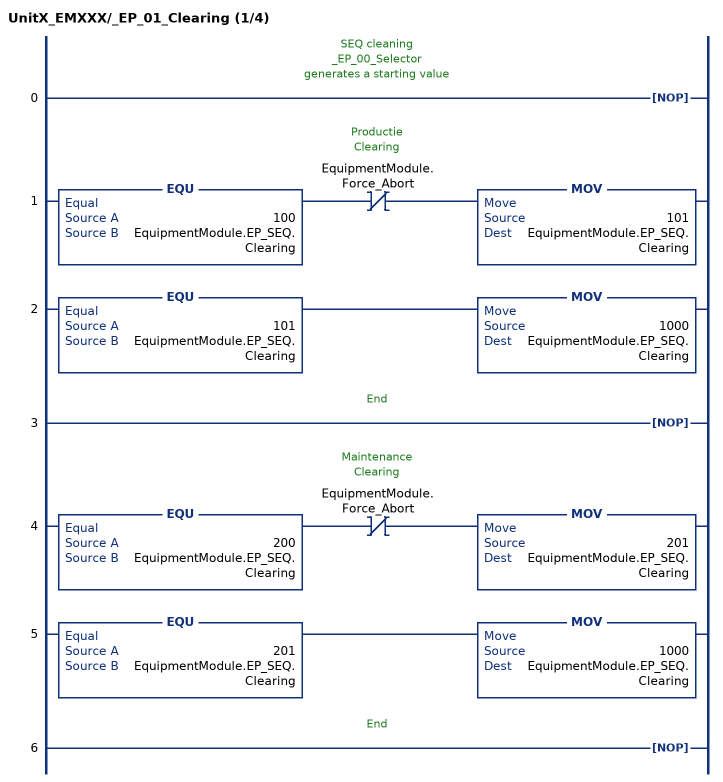
   // SEQ cleaning
   // _EP_00_Selector
   // generates a starting value
   0: NOP();
   // Productie
   // Clearing
   1: EQU(100,EquipmentModule.EP_SEQ.Clearing)XIO(EquipmentModule.Force_Abort)MOV(101,EquipmentModule.EP_SEQ.Clearing);
   2: EQU(101,EquipmentModule.EP_SEQ.Clearing)MOV(1000,EquipmentModule.EP_SEQ.Clearing);
   // End
   3: NOP();
   // Maintenance
   // Clearing
   4: EQU(200,EquipmentModule.EP_SEQ.Clearing)XIO(EquipmentModule.Force_Abort)MOV(201,EquipmentModule.EP_SEQ.Clearing);
   5: EQU(201,EquipmentModule.EP_SEQ.Clearing)MOV(1000,EquipmentModule.EP_SEQ.Clearing);
   // End
   6: NOP();
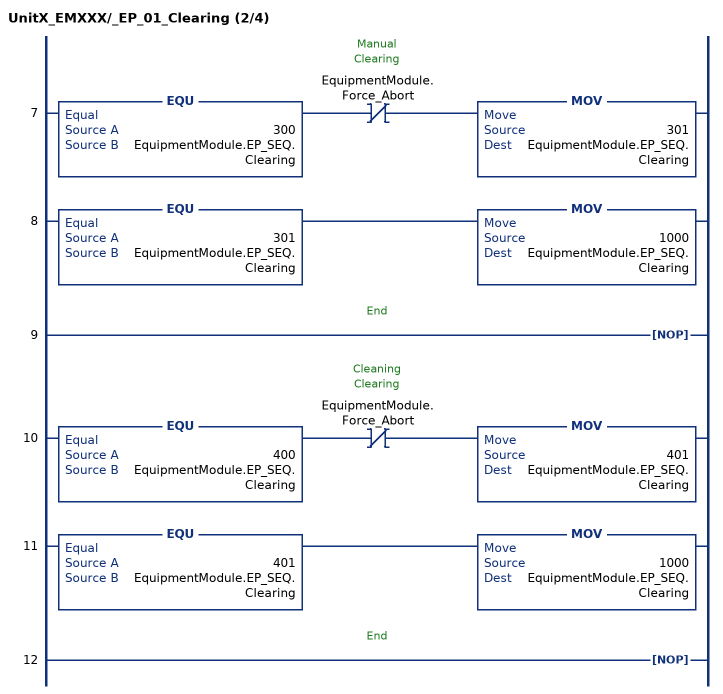
   // Manual
   // Clearing
   7: EQU(300,EquipmentModule.EP_SEQ.Clearing)XIO(EquipmentModule.Force_Abort)MOV(301,EquipmentModule.EP_SEQ.Clearing);
   8: EQU(301,EquipmentModule.EP_SEQ.Clearing)MOV(1000,EquipmentModule.EP_SEQ.Clearing);
   // End
   9: NOP();
   // Cleaning
   // Clearing
   10: EQU(400,EquipmentModule.EP_SEQ.Clearing)XIO(EquipmentModule.Force_Abort)MOV(401,EquipmentModule.EP_SEQ.Clearing);
   11: EQU(401,EquipmentModule.EP_SEQ.Clearing)MOV(1000,EquipmentModule.EP_SEQ.Clearing);
   // End
   12: NOP();
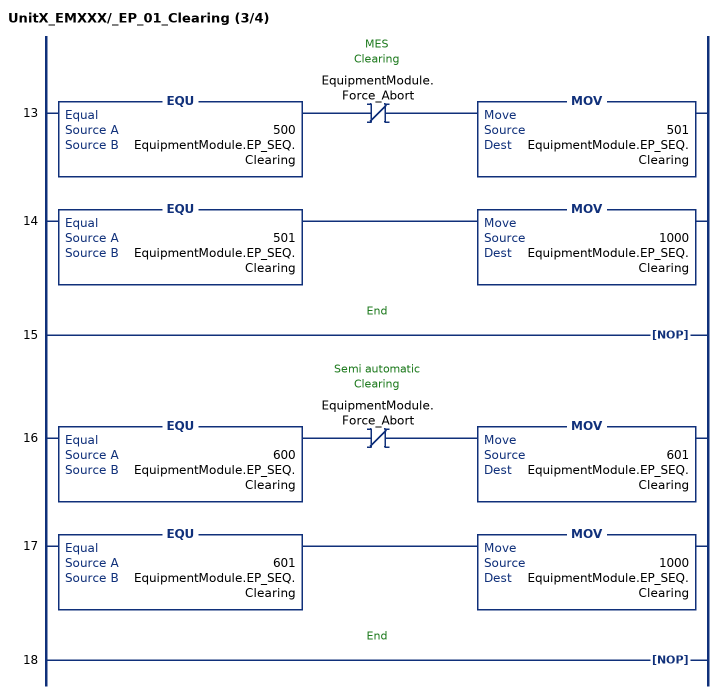
   // MES
   // Clearing
   13: EQU(500,EquipmentModule.EP_SEQ.Clearing)XIO(EquipmentModule.Force_Abort)MOV(501,EquipmentModule.EP_SEQ.Clearing);
   14: EQU(501,EquipmentModule.EP_SEQ.Clearing)MOV(1000,EquipmentModule.EP_SEQ.Clearing);
   // End
   15: NOP();
   // Semi automatic
   // Clearing
   16: EQU(600,EquipmentModule.EP_SEQ.Clearing)XIO(EquipmentModule.Force_Abort)MOV(601,EquipmentModule.EP_SEQ.Clearing);
   17: EQU(601,EquipmentModule.EP_SEQ.Clearing)MOV(1000,EquipmentModule.EP_SEQ.Clearing);
   // End
   18: NOP();
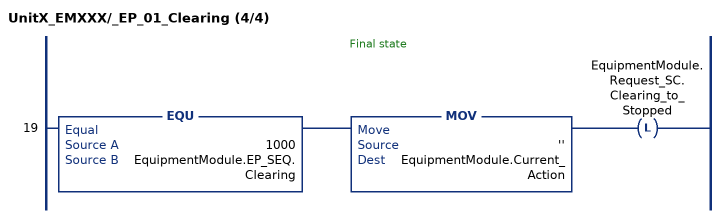
   // Final state
   19: EQU(1000,EquipmentModule.EP_SEQ.Clearing)MOV('',EquipmentModule.Current_Action)OTL(EquipmentModule.Request_SC.Clearing_to_Stopped);
END_ROUTINE

ROUTINE _EP_03_Starting   (* ladder *)
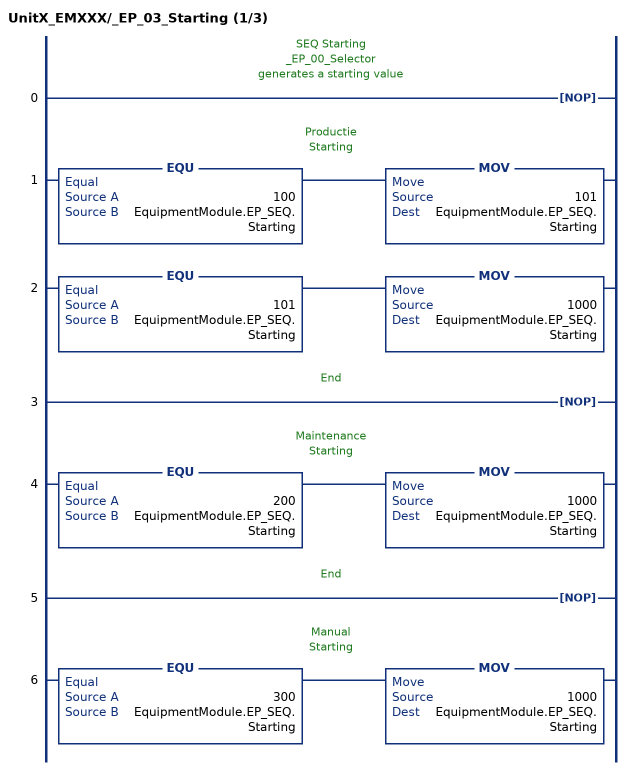
   // SEQ Starting
   // _EP_00_Selector
   // generates a starting value
   0: NOP();
   // Productie
   // Starting
   1: EQU(100,EquipmentModule.EP_SEQ.Starting)MOV(101,EquipmentModule.EP_SEQ.Starting);
   2: EQU(101,EquipmentModule.EP_SEQ.Starting)MOV(1000,EquipmentModule.EP_SEQ.Starting);
   // End
   3: NOP();
   // Maintenance
   // Starting
   4: EQU(200,EquipmentModule.EP_SEQ.Starting)MOV(1000,EquipmentModule.EP_SEQ.Starting);
   // End
   5: NOP();
   // Manual
   // Starting
   6: EQU(300,EquipmentModule.EP_SEQ.Starting)MOV(1000,EquipmentModule.EP_SEQ.Starting);
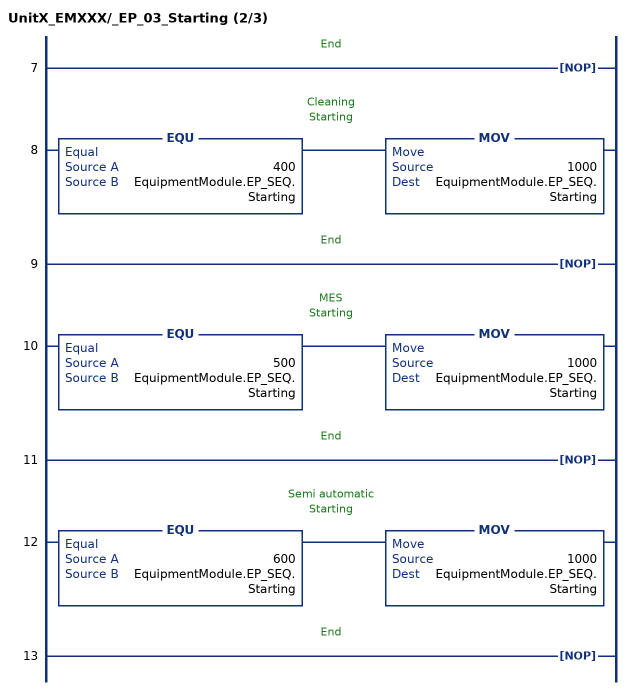
   // End
   7: NOP();
   // Cleaning
   // Starting
   8: EQU(400,EquipmentModule.EP_SEQ.Starting)MOV(1000,EquipmentModule.EP_SEQ.Starting);
   // End
   9: NOP();
   // MES
   // Starting
   10: EQU(500,EquipmentModule.EP_SEQ.Starting)MOV(1000,EquipmentModule.EP_SEQ.Starting);
   // End
   11: NOP();
   // Semi automatic
   // Starting
   12: EQU(600,EquipmentModule.EP_SEQ.Starting)MOV(1000,EquipmentModule.EP_SEQ.Starting);
   // End
   13: NOP();
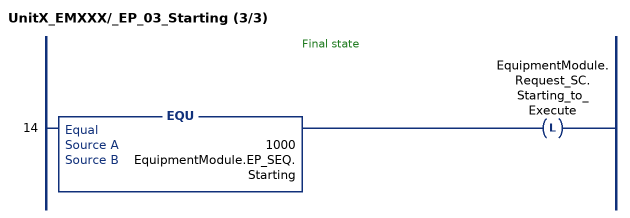
   // Final state
   14: EQU(1000,EquipmentModule.EP_SEQ.Starting)OTL(EquipmentModule.Request_SC.Starting_to_Execute);
END_ROUTINE

ROUTINE _EP_06_Execute   (* ladder *)
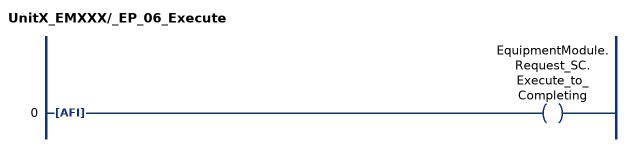
   0: AFI()OTE(EquipmentModule.Request_SC.Execute_to_Completing);
END_ROUTINE

ROUTINE _EP_07_Stopping   (* ladder *)
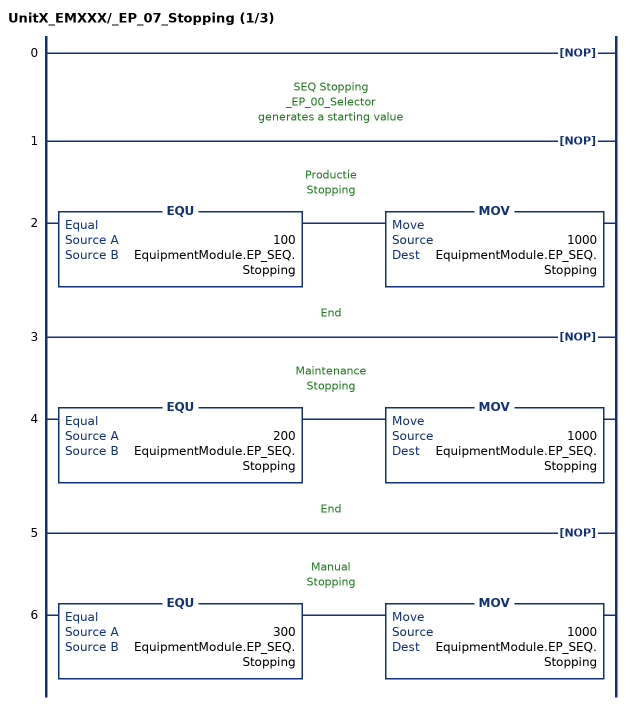
   0: NOP();
   // SEQ Stopping
   // _EP_00_Selector
   // generates a starting value
   1: NOP();
   // Productie
   // Stopping
   2: EQU(100,EquipmentModule.EP_SEQ.Stopping)MOV(1000,EquipmentModule.EP_SEQ.Stopping);
   // End
   3: NOP();
   // Maintenance
   // Stopping
   4: EQU(200,EquipmentModule.EP_SEQ.Stopping)MOV(1000,EquipmentModule.EP_SEQ.Stopping);
   // End
   5: NOP();
   // Manual
   // Stopping
   6: EQU(300,EquipmentModule.EP_SEQ.Stopping)MOV(1000,EquipmentModule.EP_SEQ.Stopping);
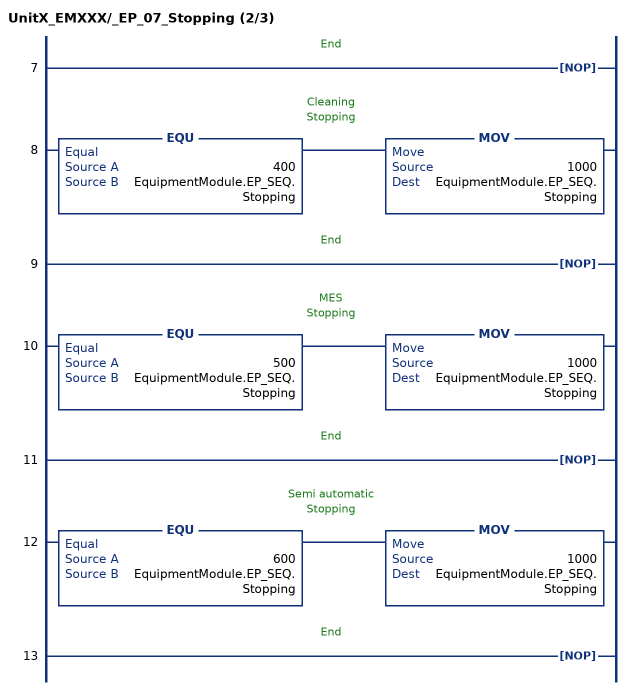
   // End
   7: NOP();
   // Cleaning
   // Stopping
   8: EQU(400,EquipmentModule.EP_SEQ.Stopping)MOV(1000,EquipmentModule.EP_SEQ.Stopping);
   // End
   9: NOP();
   // MES
   // Stopping
   10: EQU(500,EquipmentModule.EP_SEQ.Stopping)MOV(1000,EquipmentModule.EP_SEQ.Stopping);
   // End
   11: NOP();
   // Semi automatic
   // Stopping
   12: EQU(600,EquipmentModule.EP_SEQ.Stopping)MOV(1000,EquipmentModule.EP_SEQ.Stopping);
   // End
   13: NOP();
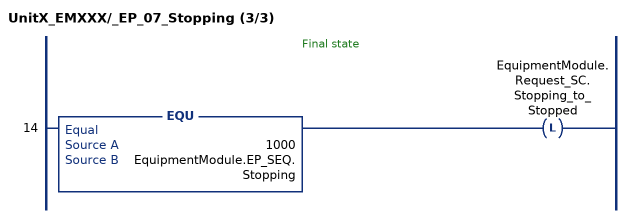
   // Final state
   14: EQU(1000,EquipmentModule.EP_SEQ.Stopping)OTL(EquipmentModule.Request_SC.Stopping_to_Stopped);
END_ROUTINE

ROUTINE _EP_08_Aborting   (* ladder *)
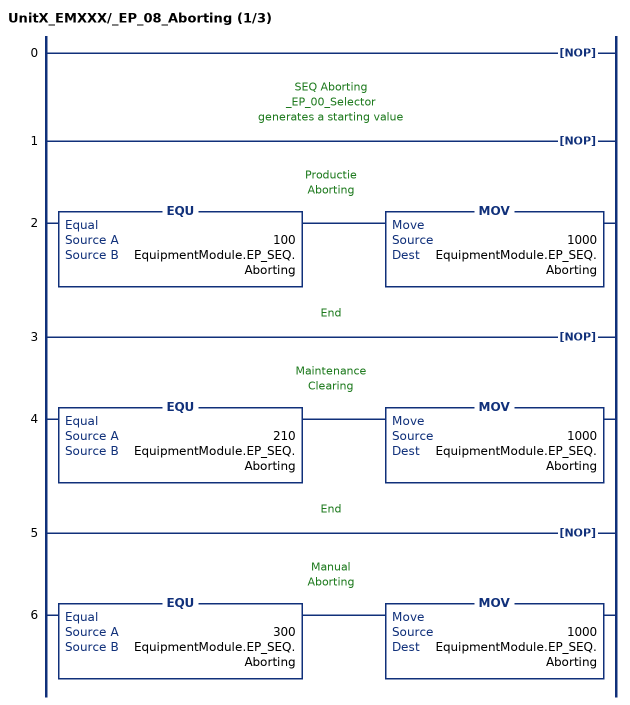
   0: NOP();
   // SEQ Aborting
   // _EP_00_Selector
   // generates a starting value
   1: NOP();
   // Productie
   // Aborting
   2: EQU(100,EquipmentModule.EP_SEQ.Aborting)MOV(1000,EquipmentModule.EP_SEQ.Aborting);
   // End
   3: NOP();
   // Maintenance
   // Clearing
   4: EQU(210,EquipmentModule.EP_SEQ.Aborting)MOV(1000,EquipmentModule.EP_SEQ.Aborting);
   // End
   5: NOP();
   // Manual
   // Aborting
   6: EQU(300,EquipmentModule.EP_SEQ.Aborting)MOV(1000,EquipmentModule.EP_SEQ.Aborting);
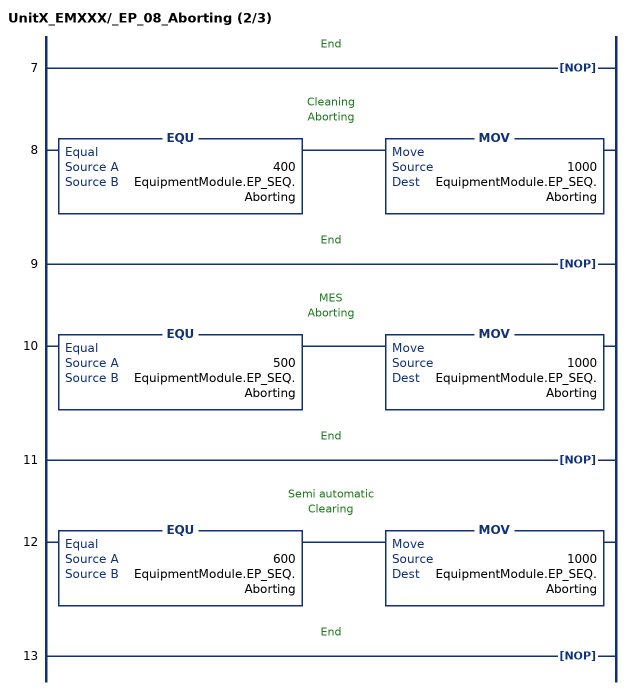
   // End
   7: NOP();
   // Cleaning
   // Aborting
   8: EQU(400,EquipmentModule.EP_SEQ.Aborting)MOV(1000,EquipmentModule.EP_SEQ.Aborting);
   // End
   9: NOP();
   // MES
   // Aborting
   10: EQU(500,EquipmentModule.EP_SEQ.Aborting)MOV(1000,EquipmentModule.EP_SEQ.Aborting);
   // End
   11: NOP();
   // Semi automatic
   // Clearing
   12: EQU(600,EquipmentModule.EP_SEQ.Aborting)MOV(1000,EquipmentModule.EP_SEQ.Aborting);
   // End
   13: NOP();
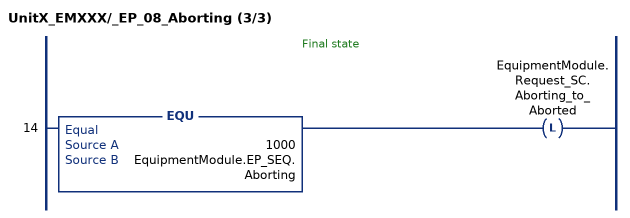
   // Final state
   14: EQU(1000,EquipmentModule.EP_SEQ.Aborting)OTL(EquipmentModule.Request_SC.Aborting_to_Aborted);
END_ROUTINE

ROUTINE _EP_10_Holding   (* ladder *)
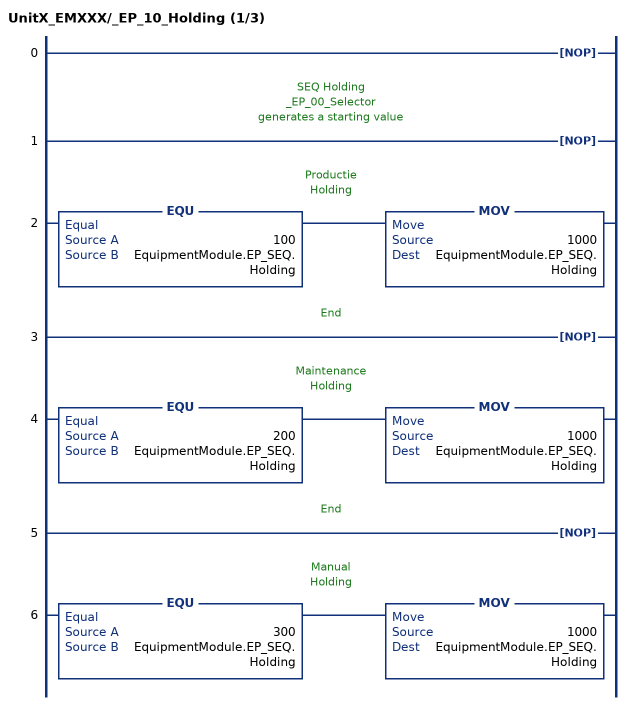
   0: NOP();
   // SEQ Holding
   // _EP_00_Selector
   // generates a starting value
   1: NOP();
   // Productie
   // Holding
   2: EQU(100,EquipmentModule.EP_SEQ.Holding)MOV(1000,EquipmentModule.EP_SEQ.Holding);
   // End
   3: NOP();
   // Maintenance
   // Holding
   4: EQU(200,EquipmentModule.EP_SEQ.Holding)MOV(1000,EquipmentModule.EP_SEQ.Holding);
   // End
   5: NOP();
   // Manual
   // Holding
   6: EQU(300,EquipmentModule.EP_SEQ.Holding)MOV(1000,EquipmentModule.EP_SEQ.Holding);
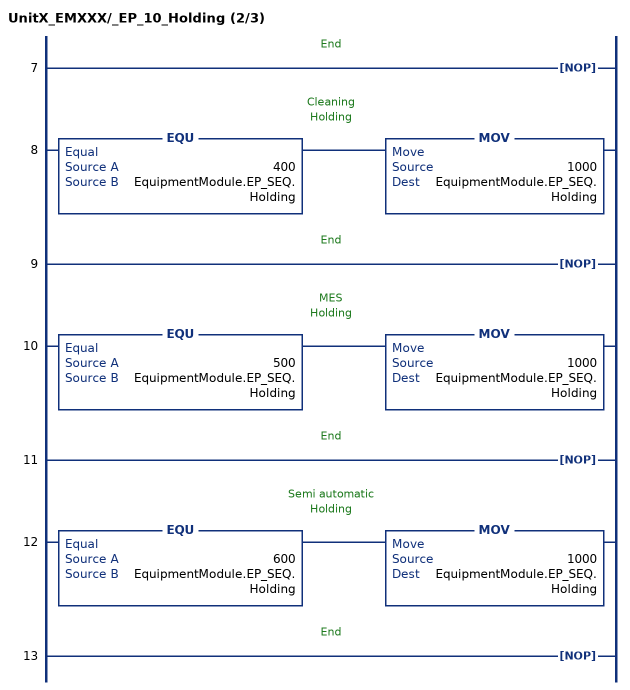
   // End
   7: NOP();
   // Cleaning
   // Holding
   8: EQU(400,EquipmentModule.EP_SEQ.Holding)MOV(1000,EquipmentModule.EP_SEQ.Holding);
   // End
   9: NOP();
   // MES
   // Holding
   10: EQU(500,EquipmentModule.EP_SEQ.Holding)MOV(1000,EquipmentModule.EP_SEQ.Holding);
   // End
   11: NOP();
   // Semi automatic
   // Holding
   12: EQU(600,EquipmentModule.EP_SEQ.Holding)MOV(1000,EquipmentModule.EP_SEQ.Holding);
   // End
   13: NOP();
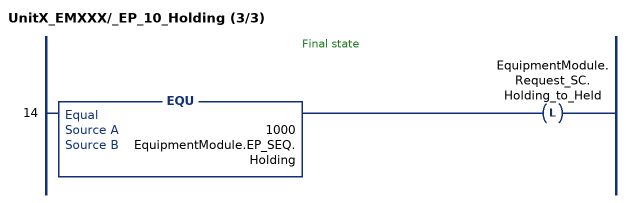
   // Final state
   14: EQU(1000,EquipmentModule.EP_SEQ.Holding)OTL(EquipmentModule.Request_SC.Holding_to_Held);
END_ROUTINE
